screen "参数修改画面" 1280x733, template "模板_2"
   on GenerateScreen: function_b456aad1(1, N); SetTag("变量_100", 17)
   TextField "文本域_7" at 30,0 size 574x42; Text '出现保养提示，请在 查看 / 유지보수 알림이 표시되면, 에서 확인하세요.'
      Visibility <- "VBS_maintenanceWarnStatus_index"
   Button "按钮_4" at 326,0 size 140x42; TextOff '自动画面 / 自動画面: / 자동화면'
      on Press: ActivateScreen("自动画面", 0)
      Visibility <- "VBS_maintenanceWarnStatus_index"
   TextField "文本域_8" at 30,0 size 714x42; Text '保养提示已隐藏，请在 查看 / 유지보수 알림 이미 숨김 , 에서 확인하세요.'
      Visibility <- "VBS_alwaysFalse"
   Button "按钮_3" at 352,0 size 168x42; TextOff '自动画面 / 自動画面: / 자동화면'
      on Press: ActivateScreen("自动画面", 0)
      Visibility <- "VBS_alwaysFalse"
   IOField "IO Field_1" at 195,85 size 121x40; FormatPattern 999
      ProcessValue <- "ST_HMI_Var_HMI_r64NianDu_QianShen_Best"
   TextField "Text Field_13" at 328,155 size 70x32; Text 'mm/s'
   IOField "IO Field_7" at 195,151 size 121x40; FormatPattern 9999
      ProcessValue <- "ST_HMI_Var_HMI_r64Velocity_ChuChe"
   TextField "Text Field_4" at 21,157 size 170x31; Text '出车速度: / 出機速度: / 외진속도:'
   TextField "Text Field_3" at 15,85 size 176x38; Text '牵伸捻度匹配值: ドラフト撚数マッチン グ値: 트위스트 연도 매칭값:'
   TextField "Text Field_9" at 21,216 size 170x38; Text '追捻开始捻度: 追撚開始撚数: 헤드 트위스트 시작 연도:'
   IOField "IO Field_4" at 195,216 size 121x40; FormatPattern 9999
      ProcessValue <- "ST_HMI_Var_HMI_r64NianDu_1"
      ObjectEnable <- "ST_HMI_Var_HMI_boNianDu_3"
   TextField "Text Field_10" at 328,220 size 70x32; Text 'T/M'
   TextField "Text Field_11" at 328,285 size 70x32; Text 'r/min'
   IOField "IO Field_5" at 195,282 size 121x40; FormatPattern 99999
      ProcessValue <- "ST_HMI_Var_HMI_r64NianSu_2"
   TextField "Text Field_24" at 15,282 size 176x38; Text '追捻锭子速度: 追撚スピンドル回転数: 헤드 트위스트 스핀들 속도:'
   TextField "Text Field_29" at 392,25 size 94x30; Text '支数: / 番手: / 번수:'
   IOField "IO Field_18" at 488,20 size 121x40; FormatPattern 99.9
      ProcessValue <- "ST_HMI_Var_HMI_r64ZhiShu_ChengSha"
   TextField "Text Field_2" at 21,25 size 170x31; Text '总捻度: / 総撚数: / 전체 연도:'
   TextField "Text Field_6" at 328,25 size 70x32; Text 'T/M'
   IOField "IO Field_43" at 195,20 size 121x40; FormatPattern 9999
      ProcessValue <- "ST_HMI_Var_HMI_r64NianDu_all"
   TextField "Text Field_7" at 615,23 size 60x32; Text 'Nm'
   Button "按钮_2" at 374,441 size 169x69; TextOn '启用按下 / 使用 / 작동 클릭:'; TextOff '启用 / 使用 / 사용'
      on Press: function_bbf3fe93(1, N)
      on Change: SetBit("ST_Calculation_Var_HMI_bo_Calculation_0_Start"); SetTag("ST_Calculation_Var_g_i16_Calculation_0_3_Select_Status", 1)
      on Release: SetBit("ST_Calculation_Var_HMI_bo_Calculation_0_Start"); SetTag("ST_Calculation_Var_g_i16_Calculation_0_3_Select_Status", 1)
   TextField "Text Field_15" at 615,155 size 60x32; Text 'r/min'
   IOField "IO Field_2" at 488,151 size 121x40; FormatPattern 99999
      ProcessValue <- "ST_HMI_Var_HMI_r64NianSu_Max"
      Appearance <- "ST_HMI_Var_HMI_boAlarm_NianDu_Time"
   IOField "IO Field_13" at 488,85 size 121x40; FormatPattern 99.9
      ProcessValue <- "ST_HMI_Var_HMI_r64Time_JiaNian"
      Appearance <- "ST_HMI_Var_HMI_boAlarm_NianDu_Time"
   TextField "Text Field_48" at 615,89 size 52x32; Text 's'
   Button "按钮_5" at 374,594 size 169x69; TextOn '返回 / リターン / 리턴'; TextOff '返回 / リターン / 리턴'
      on Release: ActivateScreen("设置画面", 0)
   Button "按钮_1" at 1106,176 size 145x54; TextOff '返回 / リターン / 리턴'
      on Click: ActivateScreen("设置画面", 0)
   TextField "Text Field_16" at 690,20 size 142x38; Text '捻缩捻度: ジャッキング．イン 開始撚数: 연축거리:'
   TextField "Text Field_20" at 690,85 size 142x38; Text '捻缩距离: ジャッキング．イン 距離: 연축 트위스트:'
   TextField "Text Field_17" at 970,24 size 63x32; Text 'T/M'
   TextField "Text Field_33" at 970,89 size 63x32; Text 'mm'
   IOField "IO Field_3" at 839,20 size 121x40; FormatPattern 9999
      ProcessValue <- "ST_HMI_Var_HMI_r64NianDu_NianSuo"
   IOField "IO Field_6" at 839,85 size 121x40; FormatPattern 999
      ProcessValue <- "ST_HMI_Var_HMI_r64Position_NianSuo"
      Appearance <- "ST_HMI_Var_HMI_boAlarm_NianSuo_PosNon"
   Button "OBJECT_107" at 400,216 size 232x40; TextOn '追捻启用 / 追撚使用 / 헤드 트위스트 사용'; TextOff '追捻启用 / EXIT / 追撚使用 / 헤드 트위스트 사용'
      on Release: SetBit("ST_HMI_Var_HMI_boNianDu_3")
      Appearance <- "ST_HMI_Var_HMI_boNianDu_3"
   Button "OBJECT_1" at 400,280 size 232x40; TextOn '追捻停用 / 追撚停止 / 헤드 트위스트 사용중지'; TextOff '追捻停用 / EXIT / 追撚停止 / 헤드 트위스트 사용중지'
      on Release: ResetBit("ST_HMI_Var_HMI_boNianDu_3"); SetTag("ST_HMI_Var_HMI_r64NianDu_1", "ST_HMI_Var_HMI_r64NianDu_all")
      Appearance <- "ST_HMI_Var_HMI_boNianDu_3"
   TextField "Text Field_34" at 970,154 size 63x33; Text 's'
   TextField "Text Field_18" at 392,85 size 94x38; Text '加捻时间: / 撚掛時間: / 연사시간:'
   TextField "Text Field_19" at 392,151 size 94x38; Text '锭子速度: スピンドル 回転数: 스핀들속도:'
   Button "按钮_6" at 672,440 size 169x69; TextOn '启用按下 / 使用 / 작동 클릭:'; TextOff '启用 / 使用 / 사용'; TextList "g_i16_Calculation_0_Status"
      Appearance <- "ST_Calculation_Var_g_i16_Calculation_0_Status"
      ProcessValue <- "ST_Calculation_Var_g_i16_Calculation_0_Status"
   TextField "Text Field_14" at 600,533 size 170x31; Text '生效总捻度: / 総撚数: / 전체 연도:'
   TextField "Text Field_23" at 600,600 size 170x31; Text '生效支数: / 総撚数: / 전체 연도:'
   TextField "Text Field_1" at 40,392 size 256x32; Text '更改参数步骤： / パラメーター変更手順: / 매개변수 변경 순서:'
   TextField "Text Field_8" at 38,445 size 277x32; Text '1.更改参数 / １．パラメーター変更 / 1.매개변수 변경'
   TextField "Text Field_12" at 38,510 size 277x32; Text '2.点击“启用” / ２．「使用」をクリック / 2.“사용”을 클릭'
   TextField "Text Field_5" at 38,575 size 277x32; Text '3.点击“返回” / ３．「リターン」をクリック / 3.리턴을 클릭'
   TextField "Text Field_21" at 695,150 size 137x38; Text '捻缩时间: ジャッキング．イン 時間: 연축시간:'
   TextField "Text Field_22" at 695,215 size 137x38; Text '捻缩速度: ジャッキング．イン 速度: 연축속도:'
   TextField "Text Field_31" at 695,285 size 137x32; Text '卷绕长度: / 巻取長: / 와인딩 길이:'
   TextField "Text Field_35" at 970,219 size 63x32; Text 'mm/s'
   TextField "Text Field_36" at 970,285 size 63x32; Text 'mm'
   IOField "IO Field_11" at 839,150 size 121x40; FormatPattern 99.9
      ProcessValue <- "ST_HMI_Var_HMI_r64Time_NianSuo"
   IOField "IO Field_12" at 839,215 size 121x40; FormatPattern 99.9
      ProcessValue <- "ST_HMI_Var_HMI_r64Velocity_NianSuo"
      Appearance <- "ST_HMI_Var_HMI_boAlarm_NianSuo_SuDuOver"
   IOField "IO Field_19" at 839,281 size 121x40; FormatPattern 9999
      ProcessValue <- "ST_HMI_Var_HMI_r64Length_JuanRao"
   IOField "IO Field_8" at 784,600 size 121x40; FormatPattern 99.9
      ProcessValue <- "ST_1TCP_g_myStructSend__lreal_20"
   IOField "IO Field_9" at 784,528 size 121x40; FormatPattern 9999
      ProcessValue <- "ST_1TCP_g_myStructSend__lreal_1"

screen "配方保存画面" 1280x733, template "模板_2"
   on GenerateScreen: function_b456aad1(1, N); SetTag("变量_100", 19)
   TextField "文本域_7" at 30,0 size 574x42; Text '出现保养提示，请在 查看 / 유지보수 알림이 표시되면, 에서 확인하세요.'
      Visibility <- "VBS_maintenanceWarnStatus_index"
   Button "按钮_4" at 326,0 size 140x42; TextOff '自动画面 / 自動画面 / 자동화면'
      on Press: ActivateScreen("自动画面", 0)
      Visibility <- "VBS_maintenanceWarnStatus_index"
   TextField "文本域_8" at 30,0 size 574x42; Text '保养提示已隐藏，请在 查看 / 유지보수 알림 이미 숨김 , 에서 확인하세요.'
      Visibility <- "VBS_alwaysFalse"
   Button "按钮_3" at 352,0 size 168x42; TextOff '自动画面 / 自動画面 / 자동화면'
      on Press: ActivateScreen("自动画面", 0)
      Visibility <- "VBS_alwaysFalse"
   IOField "IO Field_1" at 198,85 size 121x40; FormatPattern 999
      on OnFinishInput: SetBit("ST_Calculation_Var_HMI_bo_Calculation_0_Start"); SetTag("ST_Calculation_Var_g_i16_Calculation_0_3_Select_Status", 1)
      ProcessValue <- "ST_HMI_Var_HMI_r64NianDu_QianShen_Best"
   TextField "Text Field_13" at 331,155 size 70x32; Text 'mm/s'
   IOField "IO Field_7" at 198,151 size 121x40; FormatPattern 9999
      on OnFinishInput: SetBit("ST_Calculation_Var_HMI_bo_Calculation_0_Start"); SetTag("ST_Calculation_Var_g_i16_Calculation_0_3_Select_Status", 1)
      ProcessValue <- "ST_HMI_Var_HMI_r64Velocity_ChuChe"
   TextField "Text Field_4" at 24,157 size 170x31; Text '出车速度: / 出機速度: / 외진속도:'
   TextField "Text Field_3" at 18,85 size 176x38; Text '牵伸捻度匹配值: ドラフト撚数マッチン グ値: 트위스트 연도 매칭값:'
   TextField "Text Field_9" at 24,216 size 170x38; Text '追捻开始捻度: 追撚開始撚数: 헤드 트위스트 시작 연도:'
   IOField "IO Field_4" at 198,216 size 121x40; FormatPattern 9999
      on OnFinishInput: SetBit("ST_Calculation_Var_HMI_bo_Calculation_0_Start"); SetTag("ST_Calculation_Var_g_i16_Calculation_0_3_Select_Status", 1)
      ProcessValue <- "ST_HMI_Var_HMI_r64NianDu_1"
      ObjectEnable <- "ST_HMI_Var_HMI_boNianDu_3"
   TextField "Text Field_10" at 331,220 size 70x32; Text 'T/M'
   TextField "Text Field_11" at 331,285 size 70x32; Text 'r/min'
   IOField "IO Field_5" at 198,282 size 121x40; FormatPattern 99999
      on OnFinishInput: SetBit("ST_Calculation_Var_HMI_bo_Calculation_0_Start"); SetTag("ST_Calculation_Var_g_i16_Calculation_0_3_Select_Status", 1)
      ProcessValue <- "ST_HMI_Var_HMI_r64NianSu_2"
   TextField "Text Field_24" at 18,282 size 176x38; Text '追捻锭子速度: 追撚スピンドル回転数: 헤드 트위스트 스핀들 속도:'
   TextField "Text Field_29" at 366,25 size 101x30; Text '支数: / 番手: / 번수:'
   IOField "IO Field_18" at 469,20 size 121x40; FormatPattern 99.9
      ProcessValue <- "ST_HMI_Var_HMI_r64ZhiShu_ChengSha"
   TextField "Text Field_2" at 24,25 size 170x31; Text '总捻度: / 総撚数: / 전체 연도:'
   TextField "Text Field_6" at 331,25 size 70x32; Text 'T/M'
   IOField "IO Field_43" at 198,20 size 121x40; FormatPattern 9999
      on OnFinishInput: SetBit("ST_Calculation_Var_HMI_bo_Calculation_0_Start"); SetTag("ST_Calculation_Var_g_i16_Calculation_0_3_Select_Status", 1)
      ProcessValue <- "ST_HMI_Var_HMI_r64NianDu_all"
   TextField "Text Field_7" at 596,23 size 60x32; Text 'Nm'
   Button "按钮_5" at 1067,584 size 169x69; TextOff '删除数据记录 / 保存データの削除 / 데이터 기록 삭제'
      on Click: function_be763222("配方视图_1")
   Button "按钮_1" at 680,584 size 169x69; TextOff '当前值显示 / 目前値表示 / 현재값 표시'
      on Click: function_b9843780("配方视图_1")
   Button "按钮_7" at 1107,191 size 145x54; TextOff '返回 / リターン / 리턴'
      on Click: ActivateScreen("设置画面", 0)
   Button "按钮_2" at 861,584 size 193x69; TextOff '数据记录另存为 データを新たに保存する 데이터 기록을 다른 이름으로 저장'
      on Click: function_f5cdec3f("配方视图_1")
   IOField "IO Field_3" at 839,20 size 121x40; FormatPattern 9999
      ProcessValue <- "ST_HMI_Var_HMI_r64NianDu_NianSuo"
   IOField "IO Field_6" at 839,85 size 121x40; FormatPattern 999
      ProcessValue <- "ST_HMI_Var_HMI_r64Position_NianSuo"
   Button "OBJECT_107" at 400,216 size 232x40; TextOn '追捻启用 / 追撚使用 / 헤드 트위스트 사용'; TextOff '追捻启用 / EXIT / 追撚使用 / 헤드 트위스트 사용'
      on Release: SetBit("ST_HMI_Var_HMI_boNianDu_3")
      on Change: SetBit("ST_Calculation_Var_HMI_bo_Calculation_0_Start"); SetTag("ST_Calculation_Var_g_i16_Calculation_0_3_Select_Status", 1)
      Appearance <- "ST_HMI_Var_HMI_boNianDu_3"
   Button "OBJECT_1" at 400,280 size 232x40; TextOn '追捻停用 / 追撚停止 / 헤드 트위스트 사용중지'; TextOff '追捻停用 / EXIT / 追撚停止 / 헤드 트위스트 사용중지'
      on Release: ResetBit("ST_HMI_Var_HMI_boNianDu_3"); SetTag("ST_HMI_Var_HMI_r64NianDu_1", "ST_HMI_Var_HMI_r64NianDu_all")
      on Change: SetBit("ST_Calculation_Var_HMI_bo_Calculation_0_Start"); SetTag("ST_Calculation_Var_g_i16_Calculation_0_3_Select_Status", 1)
      Appearance <- "ST_HMI_Var_HMI_boNianDu_3"
   RecipeView "配方视图_1" at 681,376 size 555x188; DataRecordNrCaption '编号: / Nr.: / No.: / N.º: / N°: / 番号: / 번호: / Nr. / №:'; RecipeNameCaption '配方组名称： / Recipe Name: / レシピグループ名称: / 래서피 이름: / Reseptnavn: / Имя рецепта:'; DataRecordNameCaption '子配方名称： / Datensatzname: / Data Record Name: / Nombre de registro: / Nom d'enregistrement : / Nome del set di dati: / レシピ名称: / 데이터 레코드 이름: / Datapostnavn: / Имя блока данных:'
   TextField "Text Field_1" at 26,389 size 235x32; Text '配方保存步骤： / レシピ保存手順: / 레시피 저장 순서:'
   TextField "Text Field_8" at 23,495 size 609x32; Text '2.点击“当前值显示” / ２．「目前値表示」をクリックする / 2.“현재값 표시”를 클릭'
   TextField "Text Field_12" at 23,435 size 609x32; Text '1.选择“配方组名称” / １．「レシピグループ名称」を選択する / 1.“레시피 그룹 명칭”을 선택'
   TextField "Text Field_14" at 23,556 size 609x32; Text '3.点击“数据记录另存为” / ３．「データを新たに保存する」を選択する / 3.“데이터 기록을 다른 이름으로 저장”을 클릭'
   TextField "Text Field_15" at 23,617 size 609x63; Text '4.输入数据记录名：格式为“序号-捻度-支数-年年月月日日” ４．データ名を入力： 順番ー撚数ー番手ー年 月 日 4.데이터 기록명칭을 입력:양식은“순번-연도-번수-년년월월 일일”.'
   TextField "Text Field_16" at 97,663 size 609x32; Text '例：“01-590-265-20160811” / 例：「01－590－265－20160811」 / 예시：“01-590-265-20160811”'
   TextField "Text Field_5" at 690,20 size 142x38; Text '捻缩捻度: ジャッキング．イン 開始撚数: 연축속도:'
   TextField "Text Field_17" at 970,24 size 63x32; Text 'T/M'
   TextField "Text Field_20" at 690,85 size 142x38; Text '捻缩距离: ジャッキング．イン 距離: 연축거리:'
   TextField "Text Field_33" at 970,89 size 63x32; Text 'mm'

screen "配方选择画面" 1280x733, template "模板_2"
   on GenerateScreen: SetTag("变量_100", 18)
   TextField "文本域_7" at 30,0 size 574x42; Text '出现保养提示，请在 查看 / 유지보수 알림이 표시되면, 에서 확인하세요.'
      Visibility <- "VBS_maintenanceWarnStatus_index"
   Button "按钮_4" at 326,0 size 140x42; TextOff '自动画面 / 自動画面 / 자동화면'
      on Press: ActivateScreen("自动画面", 0)
      Visibility <- "VBS_maintenanceWarnStatus_index"
   TextField "文本域_8" at 30,0 size 574x42; Text '保养提示已隐藏，请在 查看 / 유지보수 알림 이미 숨김 , 에서 확인하세요.'
      Visibility <- "VBS_alwaysFalse"
   Button "按钮_3" at 352,0 size 168x42; TextOff '自动画面 / 自動画面 / 자동화면'
      on Press: ActivateScreen("自动画面", 0)
      Visibility <- "VBS_alwaysFalse"
   IOField "IO Field_1" at 204,85 size 121x40; FormatPattern 999
      on OnFinishInput: SetBit("ST_Calculation_Var_HMI_bo_Calculation_0_Start"); SetTag("ST_Calculation_Var_g_i16_Calculation_0_3_Select_Status", 1)
      ProcessValue <- "ST_HMI_Var_HMI_r64NianDu_QianShen_Best"
   TextField "Text Field_13" at 337,155 size 70x32; Text 'mm/s'
   IOField "IO Field_7" at 204,151 size 121x40; FormatPattern 9999
      on OnFinishInput: SetBit("ST_Calculation_Var_HMI_bo_Calculation_0_Start"); SetTag("ST_Calculation_Var_g_i16_Calculation_0_3_Select_Status", 1)
      ProcessValue <- "ST_HMI_Var_HMI_r64Velocity_ChuChe"
   TextField "Text Field_4" at 24,157 size 176x31; Text '出车速度: / 出機速度: / 외진속도:'
   TextField "Text Field_3" at 24,91 size 176x38; Text '牵伸捻度匹配值: ドラフト撚数マッチン グ値: 트위스트 연도 매칭값:'
   TextField "Text Field_9" at 24,216 size 176x38; Text '追捻开始捻度: 追撚開始撚数: 헤드 트위스트 시작 연도:'
   IOField "IO Field_4" at 204,216 size 121x40; FormatPattern 9999
      on OnFinishInput: SetBit("ST_Calculation_Var_HMI_bo_Calculation_0_Start"); SetTag("ST_Calculation_Var_g_i16_Calculation_0_3_Select_Status", 1)
      ProcessValue <- "ST_HMI_Var_HMI_r64NianDu_1"
   TextField "Text Field_10" at 337,220 size 70x32; Text 'T/M'
   TextField "Text Field_11" at 337,285 size 70x32; Text 'r/min'
   IOField "IO Field_5" at 204,282 size 121x40; FormatPattern 99999
      on OnFinishInput: SetBit("ST_Calculation_Var_HMI_bo_Calculation_0_Start"); SetTag("ST_Calculation_Var_g_i16_Calculation_0_3_Select_Status", 1)
      ProcessValue <- "ST_HMI_Var_HMI_r64NianSu_2"
   TextField "Text Field_24" at 24,282 size 176x38; Text '追捻锭子速度: 追撚スピンドル回転数: 헤드 트위스트 스핀들 속도:'
   TextField "Text Field_29" at 384,25 size 82x30; Text '支数: / 番手: / 번수:'
   IOField "IO Field_18" at 468,20 size 121x40; FormatPattern 99.9
      ProcessValue <- "ST_HMI_Var_HMI_r64ZhiShu_ChengSha"
   TextField "Text Field_2" at 24,25 size 176x31; Text '总捻度: / 総撚数 / 전체 연도:'
   TextField "Text Field_6" at 337,25 size 70x32; Text 'T/M'
   IOField "IO Field_43" at 204,20 size 121x40; FormatPattern 9999
      on OnFinishInput: SetBit("ST_Calculation_Var_HMI_bo_Calculation_0_Start"); SetTag("ST_Calculation_Var_g_i16_Calculation_0_3_Select_Status", 1)
      ProcessValue <- "ST_HMI_Var_HMI_r64NianDu_all"
   TextField "Text Field_7" at 595,23 size 60x32; Text 'Nm'
   Button "按钮_1" at 681,580 size 169x69; TextOff '启用当前配方 / 目前レシピの使用 / 현재 레시피 사용'
      on Click: function_ac24277f("配方视图_1")
      on Release: SetBit("ST_Calculation_Var_HMI_bo_Calculation_0_Start"); SetTag("ST_Calculation_Var_g_i16_Calculation_0_3_Select_Status", 1)
   Button "按钮_7" at 1106,176 size 145x54; TextOff '返回 / リターン / 리턴'
      on Click: ActivateScreen("设置画面", 0)
   RecipeView "配方视图_1" at 681,376 size 555x188; DataRecordNrCaption '编号: / Nr.: / No.: / N.º: / N°: / 番号: / 번호: / Nr. / №:'; RecipeNameCaption '配方组名称： / Recipe Name: / レシピグループ名称: / 래서피 이름: / Reseptnavn: / Имя рецепта:'; DataRecordNameCaption '子配方名称： / Datensatzname: / Data Record Name: / Nombre de registro: / Nom d'enregistrement : / Nome del set di dati: / レシピ名称: / 데이터 레코드 이름: / Datapostnavn: / Имя блока данных:'
   TextField "Text Field_1" at 40,389 size 227x32; Text '配方选择步骤： / レシピ選択手順: / 레시피 선택 순서:'
   TextField "Text Field_8" at 39,495 size 592x32; Text '2.选择“子配方名称” / ２．「レシピ名称」を選択する / 2. “하위 레시비 명칭”을 선택'
   TextField "Text Field_12" at 39,435 size 592x32; Text '1.选择“配方组名称” / １．「レシピグループ名称」を選択する / 1.“레시피 그룹 명칭”을 선택'
   TextField "Text Field_14" at 39,556 size 592x32; Text '3.点击“启用当前配方” / ３．「目前レシピ使用」をクリックする / 3. “현재 레시피 사용”을 클릭한다.'
   IOField "IO Field_9" at 839,20 size 121x40; FormatPattern 9999
      on OnFinishInput: SetBit("ST_Calculation_Var_HMI_bo_Calculation_0_Start"); SetTag("ST_Calculation_Var_g_i16_Calculation_0_3_Select_Status", 1)
      ProcessValue <- "ST_HMI_Var_HMI_r64NianDu_NianSuo"
   IOField "IO Field_10" at 839,85 size 121x40; FormatPattern 999
      on OnFinishInput: SetBit("ST_Calculation_Var_HMI_bo_Calculation_0_Start")
      Appearance <- "ST_HMI_Var_HMI_boAlarm_NianSuo_PosNon"
      ProcessValue <- "ST_HMI_Var_HMI_r64Position_NianSuo"
   TextField "Text Field_5" at 698,24 size 140x38; Text '捻缩捻度: ジャッキング．イン 開始撚数: 연축 트위스트:'
   TextField "Text Field_17" at 970,24 size 63x32; Text 'T/M'
   TextField "Text Field_20" at 700,89 size 130x38; Text '捻缩距离: ジャッキング．イン 距離: 연축거리:'
   TextField "Text Field_33" at 970,89 size 63x32; Text 'mm'

screen "常用调试画面" 1280x733
   on GenerateScreen: SetTag("变量_100", 10)
   Button "HmiScreenItemData_1" at 1105,71 size 145x54; TextOn '向后 / Back / 後向き / 뒤로'; TextOff '向后 / Back / 後向き / 뒤로'
      on Release: ActivateScreen("设置画面", 0)
   IOField "IO Field_38" at 730,162 size 112x42; FormatPattern 999
      ProcessValue <- "ST_HMI_Var_HMI_r64Axis_ZouChe_Position_KongDing_12"
   IOField "IO Field_41" at 730,54 size 112x42; FormatPattern 99
      ProcessValue <- "ST_HMI_Var_HMI_r64_MaoZhou_TouShu"
   IOField "IO Field_10" at 730,108 size 112x42; FormatPattern 999.9
      ProcessValue <- "ST_HMI_Var_HMI_r64Axis_ZouChe_Position_ShengTou_Start_Position"
   IOField "IO Field_28" at 100,322 size 108x40; FormatPattern 99.99
      ProcessValue <- "ST_HMI_Var_HMI_r64_k_ZhangLi_Rate"
   IOField "IO Field_21" at 100,270 size 108x41; FormatPattern 99.99
      ProcessValue <- "ST_HMI_Var_HMI_g1_n_delt_new_0"
   IOField "IO Field_20" at 100,216 size 108x41; FormatPattern 99.99
      ProcessValue <- "ST_HMI_Var_HMI_f1_n_delt_new_0"
   IOField "IO Field_22" at 100,163 size 108x40; FormatPattern 99.99
      ProcessValue <- "ST_HMI_Var_HMI_r64Axis_1_ZhangLi_Position_JuanRao_Set_N"
   IOField "IO Field_23" at 100,109 size 108x40; FormatPattern 99.99
      ProcessValue <- "ST_HMI_Var_HMI_r64Axis_1_ZhangLi_Position_JuanRao_Set_ND"
   IOField "IO Field_24" at 100,55 size 108x40; FormatPattern 99.99
      ProcessValue <- "ST_HMI_Var_HMI_r64Axis_1_ZhangLi_Position_JuanRao_Set_0"
   IOField "IO Field_57" at 100,427 size 109x41; FormatPattern 9.99
      ProcessValue <- "ST_HMI_Var_HMI_k_TuiRao"
   IOField "IO Field_58" at 100,480 size 109x41; FormatPattern 9.99
      ProcessValue <- "ST_HMI_Var_HMI_scalevalue_Cam_3"
   IOField "IO Field_1" at 100,594 size 108x40; FormatPattern 99999
      ProcessValue <- "ST_Main_Var_g_r64Axis_DingZi_PositiveAccel_CunRao"
   IOField "IO Field_25" at 100,648 size 108x40; FormatPattern 99.99
      ProcessValue <- "ST_Main_Var_g_r64Axis_DingZi_Velocity_CunRao_ratio"
   Button "HmiScreenItemData_2" at 1104,352 size 145x54; TextOn '向后 / 後向き / 뒤로'; TextOff '张力测定 / 張力測定 / 장력 측정'; Authorization "Operate_4"
      on Release: ActivateScreen("张力测定", 0)
   Button "HmiScreenItemData_3" at 1104,424 size 145x54; TextOn '向后 / 後向き / 뒤로'; TextOff '原点设定 / 原点設定 / 원점 설정'; Authorization "Operate_4"
      on Release: ActivateScreen("原点设定", 0)
   Button "HmiScreenItemData_4" at 1104,496 size 145x54; TextOn '向后 / 後向き / 뒤로'; TextOff '纱管参数设定 糸管パラメーター 設定 보빈 매개변수 설정'; Authorization "Operate_4"
      on Release: ActivateScreen("纱管参数设定", 0)
   Button "Template_Button_1" at 791,673 size 85x59; TextOff 'Text'; PictureOff "China_1"
      on Click: function_fb9197e8(-1)
   Button "HmiScreenItemData_15" at 928,679 size 158x53; TextOn '6卷绕相关1 / 6巻取関係1'; TextOff '校准触摸屏 / タッチパネルの校正 / 터치 스크린 교정'
      on Release: function_bc3e350c()
   IOField "IO Field_2" at 729,214 size 112x42; FormatPattern 99.9
      ProcessValue <- "ST_HMI_Var_HMI_r64Axis_ZouChe_Position_ZiDongTingZhi"
   IOField "IO Field_3" at 729,270 size 112x42; FormatPattern 999
      ProcessValue <- "ST_HMI_Var_HMI_r64Axis_ZouChe_Position_ChuChe_Middle"
   Button "HmiScreenItemData_6" at 1104,570 size 145x54; TextOn '向后 / 後向き / 뒤로'; TextOff '纱穗参数设定 糸管パラメーター 設定 코프 매개변수'; Authorization "Operate_4"
      on Release: ActivateScreen("纱穗参数设定", 0)
   IOField "IO Field_8" at 728,392 size 112x42; FormatPattern 99999
      Visibility <- "ST_Calculation_Var_Date_Temp"
      ProcessValue <- "ST_Calculation_Var_g_r64Axis_DingZi_PositiveAccel_Buffer_JiaNian{1}"
      Appearance <- "ST_HMI_Var_HMI_boAlarm_NianDu_Time"
   IOField "IO Field_7" at 728,392 size 112x42; FormatPattern 99999
      Visibility <- "ST_Calculation_Var_Date_Temp"
      ProcessValue <- "ST_Calculation_Var_g_r64Axis_DingZi_PositiveAccel_Buffer_JiaNian{0}"
      Appearance <- "ST_HMI_Var_HMI_boAlarm_NianDu_Time"
   Button "Template_Button_11" at 1196,673 size 78x59; TextOn 'NavigateHome'; TextOff 'NavigateHome'; PictureOn "NavigateHome_TP1200_Comfort"; PictureOff "NavigateHome_TP1200_Comfort"
      on Release: ActivateScreen("自动画面", 0); function_f23ef4c9()
   TextField "Text Field_44" at 219,427 size 290x41; Text '退绕曲线拐点比例 / パッキングオフ湾曲点比例 / 언와인딩 곡선 변곡점 비율'
   TextField "Text Field_46" at 219,480 size 254x41; Text '退绕圈数比例 / パッキングオフ巻取比例 / 언와인딩 랩수 비율'
   TextField "Text Field_37" at 222,218 size 430x41; Text '卷绕速度中点调整值—初始值 / 中間点の取り巻き速度調整値ー初期値 / 와인딩 속도 중심점조정값-초기값'
   TextField "Text Field_38" at 222,272 size 430x41; Text '卷绕速度末点调整值—初始值 / 終了時点の取り巻き速度調整値ー初期値 / 와인딩 속도 종료점조정값-초기값'
   TextField "Text Field_39" at 222,165 size 430x41; Text '卷绕张力弓目标值—满纱时 / カウンターフォーラーの目標値ー満巻時 / 와인딩 장력 호랑 목표값-만사일시'
   TextField "Text Field_40" at 224,112 size 430x41; Text '卷绕张力弓目标值—最大直径时 / カウンターフォーラーの目標値ー最大直径時 / 와이딩 장력 호랑목표값-최대직경일시'
   TextField "Text Field_41" at 222,57 size 430x41; Text '卷绕张力弓目标值—生头时 / カウンターフォーラーの目標値ー巻始め / 와인딩 장력호랑 목표값-실시작점'
   TextField "Text Field_45" at 222,324 size 430x41; Text '卷绕张力弓反馈增益 / カウンターフォーラーのフィードバック増幅 / 와인딩 장력호랑 피드백 게인'
   TextField "Text Field_1" at 222,592 size 430x41; Text '存绕锭子加速度 / 逆巻取スピンドル加速度 / 와인딩 스핀들 가속'
   TextField "Text Field_42" at 222,646 size 430x41; Text '存绕锭子速度比例 / 逆巻取スピンドル回転速度比例 / 와인딩 스핀들 속도 비율'
   TextField "Text Field_58" at 857,164 size 230x41; Text '生头中间停止位置 / 自動停止位置 / 스레딩중 정지위치'
   TextField "Text Field_8" at 857,56 size 230x41; Text '毛轴头数 / 篠棒本数 / 시누 세부샤프트개수'
   TextField "Text Field_2" at 857,110 size 230x41; Text '生头起点位置 / 口付け開始点位置 / 스레딩시작점 위치'
   TextField "Text Field_14" at 100,6 size 233x42; Text '卷绕相关 / 巻取関係 / 와인딩 관련'
   TextField "Text Field_3" at 100,377 size 233x42; Text '退绕相关 / パッキングオフ関連 / 언와인딩 관련'
   TextField "Text Field_4" at 100,542 size 233x42; Text '存绕相关 / 逆巻取関連 / 와인딩관련'
   TextField "Text Field_5" at 778,6 size 233x42; Text '其他 / その他 / 기타'
   Button "按钮_1" at 1104,280 size 145x54; TextOff '牵伸调整 / 연신조절'; Authorization "Operate_4"
      on Press: ActivateScreen("牵伸调整画面", 0)
   TextField "Text Field_6" at 856,216 size 230x41; Text '自动停止位置 / 自動停止位置 / 자동정지위치'
   TextField "Text Field_7" at 856,272 size 230x41; Text '出车停止位置 / 自動停止位置 / 외진정지위치'
   IOField "IO Field_4" at 728,452 size 112x42; FormatPattern 9.99
      on OnFinishInput: SetBit("ST_Calculation_Var_HMI_bo_Calculation_0_Start"); SetTag("ST_Calculation_Var_g_i16_Calculation_0_3_Select_Status", 1)
      ProcessValue <- "ST_TO_DZ_FU_Var_HMI_r64Ratio_PositiveAccelStartJerk_JiaNian"
   IOField "IO Field_6" at 728,508 size 112x42; FormatPattern 9.99
      on OnFinishInput: SetBit("ST_Calculation_Var_HMI_bo_Calculation_0_Start"); SetTag("ST_Calculation_Var_g_i16_Calculation_0_3_Select_Status", 1)
      ProcessValue <- "ST_TO_DZ_FU_Var_HMI_r64Ratio_PositiveAccelEndJerk_JiaNian"
   IOField "IO Field_9" at 728,560 size 112x42; FormatPattern 99.99
      ProcessValue <- "ST_HMI_Var_HMI_r64_DingZi_Zouche_ratio_KongDing_65_1"
   TextField "Text Field_12" at 856,392 size 230x41; Text '锭子加速度'
   TextField "Text Field_9" at 856,448 size 230x41; Text '锭子+Jerk比例'
   TextField "Text Field_11" at 856,504 size 230x41; Text '锭子-Jerk比例'
   TextField "Text Field_13" at 856,560 size 230x41; Text '光锭卷绕传动比1'
   IOField "IO Field_5" at 728,320 size 112x42; FormatPattern 9.99
      on OnFinishInput: SetBit("ST_Calculation_Var_HMI_bo_Calculation_0_Start"); SetTag("ST_Calculation_Var_g_i16_Calculation_0_3_Select_Status", 1)
      ProcessValue <- "ST_HMI_Var_HMI_r64Ratio_PositiveAccel_Jerk_JiaNian"
   TextField "Text Field_10" at 856,320 size 230x41; Text '锭子加速度比例 / 自動停止位置 / 외진정지위치'
   Button "按钮_3" at 1104,208 size 145x54; TextOff '卷绕调整 / 牵伸调整 / 연신조절'; Authorization "Operate_4"
      on Press: ActivateScreen("卷绕经验参数", 0)
   Button "HmiScreenItemData_12" at 1105,138 size 146x52; TextOn '11生头相关'; TextOff '生头相关'; Authorization "Operate_4"
      on Release: ActivateScreen("生头相关", 0)
   Button "Template_Button_2" at 667,673 size 78x59; TextOff 'Text'; PictureOff "1"
      on Click: StopRuntime(0)

screen "张力测定" 1280x733, template "模板_2"
   on GenerateScreen: SetTag("变量_100", 12)
   Button "OBJECT_109" at 120,48 size 182x70; TextOn '张力测定 / 張力測定 / 장력 측정'; TextOff '张力测定 / EXIT / 張力測定 / 장력 측정'
      on Press: SetTag("ST_Main_Var_g_i16_Mode_Selected", 256)
      Appearance <- "ST_Main_Var_g_bo_Mode_Enabled_Manual"
   Button "OBJECT_110" at 120,234 size 182x70; TextOff '张力测定启动 / EXIT / 張力測定起動 / 장력 측정 시작'
      on Release: ResetBit("ST_HMI_Var_HMI_bo_ZhangLi_CeDing_Start")
      on Press: SetBit("ST_HMI_Var_HMI_bo_ZhangLi_CeDing_Start")
      Appearance <- "ST_Main_Var_g_bo_Mode_Enabled_Manual"
   IOField "I/O 域_1" at 502,42 size 86x40; FormatPattern 99.99
      ProcessValue <- "ST_Var_ZLCD_HMI_r64Axis_1_ZhangLi_Torque_CeDing_N{0}"
   IOField "I/O 域_2" at 502,86 size 86x40; FormatPattern 99.99
      ProcessValue <- "ST_Var_ZLCD_HMI_r64Axis_1_ZhangLi_Torque_CeDing_N{1}"
   IOField "I/O 域_3" at 502,130 size 86x40; FormatPattern 99.99
      ProcessValue <- "ST_Var_ZLCD_HMI_r64Axis_1_ZhangLi_Torque_CeDing_N{2}"
   IOField "I/O 域_4" at 502,174 size 86x40; FormatPattern 99.99
      ProcessValue <- "ST_Var_ZLCD_HMI_r64Axis_1_ZhangLi_Torque_CeDing_N{3}"
   IOField "I/O 域_5" at 502,218 size 86x40; FormatPattern 99.99
      ProcessValue <- "ST_Var_ZLCD_HMI_r64Axis_1_ZhangLi_Torque_CeDing_N{4}"
   IOField "I/O 域_6" at 502,261 size 86x40; FormatPattern 99.99
      ProcessValue <- "ST_Var_ZLCD_HMI_r64Axis_1_ZhangLi_Torque_CeDing_N{6}"
   Button "按钮_1" at 726,234 size 182x70; TextOn '调整 / 調整 / 조정'; TextOff '调整 / 調整 / 조정'
      on Release: ResetBit("ST_Var_ZLCD_HMI_bo_ZhangLi_CeDing_Adjustment")
      on Press: SetBit("ST_Var_ZLCD_HMI_bo_ZhangLi_CeDing_Adjustment")
   TextField "文本域_6" at 60,336 size 996x358; Text '张力弓整定步骤 1. 按一下“手动”按钮，按“成形弓降”按钮，将成形钢丝降到锭尖附近，按一下“去使能”按钮 2. 拉住张力弓，同时按住“停止”和“张力弓降”两个按钮，张力电机抱闸会松开电机抱闸，让张 力钢丝掉到走车撞块上 3. 按一下“手动按钮” 4. 点击“张力测定”，点击“张力测定启动” 5. 张力钢丝自动从最低点开始缓慢上升，同时自动记录数据 6. 待上升到48.5左右时张力弓停下 7. 观察以上6个数据，按下右侧的“调整”按钮，可看到前三个数据被第四个覆盖 8. 按下手动——>张力弓降，将张力钢丝降到正常位置 9. 结束 カウンターフォーラー調整手順 １．”手動”を一度押し、”ワイディングフォーラー下降”ボタンを押して”ワイディングフォーラー”ワイヤをスピンド ルの先端までさげ、”長期停止”ボタンを一度押す。 ２．”カウンターフォーラー”を引きながら、同時に”停止”と”カウンターフォーラー下降”ボタンを一度押す。カウ ンターモーターの制動を緩み、”ワイディングフォーラー”ワイヤをキャレージのブロックに落とせる。 ３．一度”手動”ボタンを押す ４．”張力測定”をクリックし、また”張力測定起動”をクリックする。 ５．カウンターワイヤを自動で下死点から徐々に上昇させながら、同時に自動でデータを記録する。 ６．48.5前後に上昇となった時点で、カウンターフォーラーを停止させる。 ７．以上の六つのデータを観察しながら、右側の”調整”ボタンを一度押すと、前の三つのテータが四つ目のデ ータに切り替わったことが分かる。 8．順序に”手動”と”カウンターフォーラー下降”ボタンを押せ、カウンターワイヤをさげる。 9．终。 장력 호랑셋업 순서 1. “수동”버튼을 누르고 “성형호랑하강” 버튼을 눌러 성형호랑 을스핀들 팁 근처까지 내려오게 하고 ‘비활성화’버튼을 누른다. 2. 장력호랑을당기고“정지”와 “장력호랑하강”두 버튼을 동시에 누른다.장력 호랑모터 브레이크가 풀리 면서 장력 와이어가 캐리지링크 스토퍼에 떨어진다. 3. “수동버튼”을 누른다. 4. “장력측정”을클릭하고“장력측정 시작”을 클릭한다. 5. 장력 와이어는 자동으로 최저포인트로부터 시작하여 천천히 상승하면서 자동으로 데이터를 기록한다. 6. 48. 5좌우까지 상승하면 장력 호랑을 정지한다. 7. 이상 6개데이터를 관찰하고 우측의 “조정”버튼을 누르면 처음3개 데이터가 네번째에 의해커버되어 있 는것을 볼수 있다. 8. 수동——>장력 호랑하강을 눌러 장력 와이어를 정상위치까지 내린다. 9. 종료'
   TextField "文本域_1" at 30,541 size 17x21; Text 'Text'
   Button "HmiScreenItemData_2" at 1106,174 size 145x54; TextOn '向后 / 後向き / 뒤로'; TextOff '向后 / 後向き / 뒤로'
      on Release: ActivateScreen("设置画面", 0)
   Button "HmiScreenItemData_3" at 1106,362 size 145x54; TextOn '向后 / 後向き / 뒤로'; TextOff '张力测定 / 張力測定 / 장력 측정'
      on Release: ActivateScreen("张力测定", 0)
   Button "HmiScreenItemData_4" at 1106,452 size 145x54; TextOn '向后 / 後向き / 뒤로'; TextOff '原点设定 / 原点設定 / 원점 설정'
      on Release: ActivateScreen("原点设定", 0)
   Button "HmiScreenItemData_5" at 1106,542 size 145x54; TextOn '向后 / 後向き / 뒤로'; TextOff '纱管参数设定 糸管パラメーター 設定 보빈 매개변수 설정'
      on Release: ActivateScreen("纱管参数设定", 0)
   Button "HmiScreenItemData_6" at 1106,272 size 145x54; TextOn '向后 / 後向き / 뒤로'; TextOff '常用调试画面 / 常用調整画面 / 상용 조정화면'
      on Release: ActivateScreen("常用调试画面", 0)

screen "原点设定" 1280x733, template "模板_2"
   on GenerateScreen: SetTag("变量_100", 13)
   IOField "I/O 域_1" at 885,196 size 88x48; FormatPattern 99
      ProcessValue <- "ST_HMI_Var_HMI_r64StartPosition_Axis_ZouChe_0"
   TextField "文本域_1" at 78,194 size 260x48; Text '走车编码器当前位置 キャレージのエンコー ダーの目前位置 캐리지 인코더 현재 위치'
   IOField "I/O 域_2" at 351,194 size 88x48; FormatPattern 99999.99
      ProcessValue <- "Axis_ZouChe_positioningState_actualPosition"
   Button "按钮_4" at 789,195 size 76x47; TextOff '出车 / 出機 / 외진'
      on Release: ResetBit("ST_HMI_Var_HMI_bo_ChuChe")
      on Press: SetBit("ST_HMI_Var_HMI_bo_ChuChe")
   Button "按钮_5" at 458,194 size 76x47; TextOff '进车 / 入機 / 내진'
      on Release: ResetBit("ST_HMI_Var_HMI_bo_JinChe")
      on Press: SetBit("ST_HMI_Var_HMI_bo_JinChe")
   IOField "I/O 域_3" at 885,304 size 88x48; FormatPattern 99.999
      ProcessValue <- "ST_HMI_Var_HMI_r64StartPosition_Axis_1_ZhangLi_0"
   IOField "I/O 域_4" at 885,413 size 88x48
      ProcessValue <- "ST_HMI_Var_HMI_r64StartPosition_Axis_ChengXing_0"
   TextField "文本域_2" at 78,302 size 260x48; Text '张力编码器当前位置 カウンターのエンコー ダーの目前位置 장력 인코더 현재 위치'
   IOField "I/O 域_5" at 351,302 size 88x48; FormatPattern 999.99
      ProcessValue <- "Axis_1_ZhangLi_positioningState_actualPosition"
   Button "按钮_1" at 789,303 size 76x47; TextOff '升 / 上昇 / 상승'
      on Release: ResetBit("ST_HMI_Var_HMI_bo_ZhangLi_Up")
      on Press: SetBit("ST_HMI_Var_HMI_bo_ZhangLi_Up")
   Button "按钮_2" at 458,302 size 76x47; TextOff '降 / 下降 / 하강'
      on Release: ResetBit("ST_HMI_Var_HMI_bo_ZhangLi_Down")
      on Press: SetBit("ST_HMI_Var_HMI_bo_JinChe")
   TextField "文本域_3" at 78,412 size 260x48; Text '成形编码器当前位置 ワインディングのエンコ ーダーの目前位置 성형 인코더 현재 위치'
   IOField "I/O 域_6" at 351,412 size 88x48; FormatPattern 9999.99
      ProcessValue <- "Axis_ChengXing_positioningState_actualPosition"
   Button "按钮_3" at 458,413 size 76x47; TextOff '升 / 上昇 / 상승'
      on Release: ResetBit("ST_HMI_Var_HMI_bo_ChengXing_Up")
      on Press: SetBit("ST_HMI_Var_HMI_bo_ChuChe")
   Button "按钮_6" at 789,414 size 76x47; TextOff '降 / 下降 / 하강'
      on Release: ResetBit("ST_HMI_Var_HMI_bo_ChengXing_Down")
      on Press: SetBit("ST_HMI_Var_HMI_bo_ChengXing_Down")
   Bar "棒图_1" at 554,195 size 216x49; MinimumValue 40; MaximumValue 90
      ProcessValue <- "Axis_ZouChe_positioningState_actualPosition"
   Bar "棒图_2" at 554,301 size 216x49; MinimumValue 50; MaximumValue 70
      ProcessValue <- "Axis_1_ZhangLi_positioningState_actualPosition"
   Bar "棒图_3" at 554,410 size 216x49; MinimumValue 320; MaximumValue 335
      ProcessValue <- "Axis_ChengXing_positioningState_actualPosition"
   Button "按钮_7" at 56,618 size 280x50; TextOn '微调模式 / 微調整'; TextOff '按下进入微调模式 / 微調整モードに切り替える / 미세조정 모드진입 을 누른다.'
      on Release: ResetBit("ST_HMI_Var_HMI_boMinorAdjustment_select")
      on Press: SetBit("ST_HMI_Var_HMI_boMinorAdjustment_select")
   Button "HmiScreenItemData_2" at 846,683 size 159x48; TextOn '报警画面 / 警報画面 / 경보알람화면'; TextOff '报警画面 / 警報画面 / 경보알람화면'
      on Release: ActivateScreen("报警画面", 0)
   Button "OBJECT_106" at 1039,2 size 238x42; TextOff '手动 / EXIT / 手動 / 수동'; TextList "mode_enabled_1"
      ProcessValue <- "ST_Main_Var_g_i16_Mode_Enabled"
      Appearance <- "ST_Main_Var_g_i16_Mode_Enabled"
   TextField "文本域_6" at 168,88 size 807x58; Text '注意： 不要随意修改此页的数据，不当的数据可能导致行程超限撞车的危险！ 注意：勝手に本ページのデータを変えてはいけない。不当なデータはキャレージのストロー クのオーバーを招き衝突の危険がある。 주의:임의로 이 페이지의 데이터를 수정하지 마십시오.부적절한 데이터는 스트로크 오버런충돌 위험을 초래할수 있습니다!'
   GraphicView "图形视图_2" at 57,70 size 102x99; Picture "图形_2"
   Button "HmiScreenItemData_3" at 1106,174 size 145x54; TextOn '向后 / 後向き / 뒤로'; TextOff '向后 / 後向き / 뒤로'
      on Release: ActivateScreen("设置画面", 0)
   Button "HmiScreenItemData_4" at 1106,362 size 145x54; TextOn '向后 / 後向き / 뒤로'; TextOff '张力测定 / 張力測定 / 장력 측정'
      on Release: ActivateScreen("张力测定", 0)
   Button "HmiScreenItemData_5" at 1106,452 size 145x54; TextOn '向后 / 後向き / 뒤로'; TextOff '原点设定 / 原点設定 / 원점 설정'
      on Release: ActivateScreen("原点设定", 0)
   Button "HmiScreenItemData_6" at 1105,542 size 147x54; TextOn '向后 / 後向き / 뒤로'; TextOff '纱管参数设定 糸管パラメーター 設定 보빈 매개변수 설정'
      on Release: ActivateScreen("纱管参数设定", 0)
   Button "HmiScreenItemData_7" at 1106,272 size 145x54; TextOn '向后 / 後向き / 뒤로'; TextOff '常用调试画面 / 常用調整画面 / 상용 조정화면'
      on Release: ActivateScreen("常用调试画面", 0)

screen "纱管参数设定" 1280x733, template "模板_2"
   on GenerateScreen: SetTag("变量_100", 14)
   IOField "IO Field_41" at 69,59 size 112x42; FormatPattern 99.99
      ProcessValue <- "ST_HMI_Var_HMI_r64_h0_s"
   IOField "IO Field_46" at 69,169 size 112x42; FormatPattern 99.99
      ProcessValue <- "ST_HMI_Var_HMI_r64Diameter_ShaGuan_Middle"
   IOField "IO Field_1" at 69,113 size 112x42; FormatPattern 99.99
      ProcessValue <- "ST_HMI_Var_HMI_r64Diameter_ShaGuan_Bottom"
   IOField "IO Field_2" at 69,279 size 112x42
      ProcessValue <- "ST_HMI_Var_HMI_r64Height_ShaGuan_Middle"
   IOField "IO Field_3" at 69,335 size 112x42
      ProcessValue <- "ST_HMI_Var_HMI_r64Height_ShaGuan_Top"
   IOField "IO Field_6" at 69,223 size 112x42; FormatPattern 99.99
      ProcessValue <- "ST_HMI_Var_HMI_r64Diameter_ShaGuan_Top"
   IOField "IO Field_4" at 69,392 size 112x42; FormatPattern 99.9
      ProcessValue <- "ST_HMI_Var_HMI_r64_DingZi_Zouche_ratio_KongDing_9_Shaguan1"
   IOField "IO Field_5" at 589,59 size 112x42; FormatPattern 99.99
      ProcessValue <- "ST_HMI_Var_HMI_r64_h0_s_2"
   IOField "IO Field_7" at 589,169 size 112x42; FormatPattern 99.99
      ProcessValue <- "ST_HMI_Var_HMI_r64Diameter_ShaGuan_Middle_2"
   IOField "IO Field_8" at 589,113 size 112x42; FormatPattern 99.99
      ProcessValue <- "ST_HMI_Var_HMI_r64Diameter_ShaGuan_Bottom_2"
   IOField "IO Field_9" at 589,279 size 112x42
      ProcessValue <- "ST_HMI_Var_HMI_r64Height_ShaGuan_Middle_2"
   IOField "IO Field_10" at 589,335 size 112x42
      ProcessValue <- "ST_HMI_Var_HMI_r64Height_ShaGuan_Top_2"
   IOField "IO Field_11" at 589,223 size 112x42; FormatPattern 99.99
      ProcessValue <- "ST_HMI_Var_HMI_r64Diameter_ShaGuan_Top_2"
   IOField "IO Field_12" at 589,392 size 112x42; FormatPattern 99.9
      ProcessValue <- "ST_HMI_Var_HMI_r64_DingZi_Zouche_ratio_KongDing_9_Shaguan2"
   TextField "Text Field_8" at 207,59 size 332x42; Text '纱管安装高度 / 糸管装着高度 / 보빈 설치 높이'
   TextField "Text Field_9" at 207,113 size 332x42; Text '纱管底部直径 / 糸管底部直径 / 보빈 하단부분 직경'
   TextField "Text Field_10" at 207,169 size 332x42; Text '纱管中间直径 / 糸管中間部直径 / 보빈 중간부분 직경'
   TextField "Text Field_11" at 207,223 size 332x42; Text '纱管顶部有效直径 / 糸管上部有効直径 / 보빈 상단 유효 직경'
   TextField "Text Field_12" at 207,279 size 332x42; Text '纱管从底部到中间的高度 / 糸管底部から中間部までの高度 / 보빈 하단에서 중간까지의 높이'
   TextField "Text Field_13" at 207,335 size 345x42; Text '纱管从中间到顶部的高度 / 糸管中間部から上部までの高度 / 보빈 중간부분에서 상단까지의 높이'
   TextField "Text Field_1" at 207,392 size 332x42; Text '空锭-锭子走车传动比 / 空鍾－スピンドル キャレージ伝動比 / 아이들 스핀들-스핀들 캐리지 기어비'
   TextField "Text Field_3" at 727,59 size 332x42; Text '纱管安装高度 / 糸管装着高度 / 보빈 설치 높이'
   TextField "Text Field_4" at 727,113 size 332x42; Text '纱管底部直径 / 糸管底部直径 / 보빈 하단부분 직경'
   TextField "Text Field_5" at 727,169 size 332x42; Text '纱管中间直径 / 糸管中間部直径 / 보빈 중간부분 직경'
   TextField "Text Field_6" at 727,223 size 332x42; Text '纱管顶部有效直径 / 糸管上部有効直径 / 보빈 상단 유효 직경'
   TextField "Text Field_7" at 727,279 size 332x42; Text '纱管从底部到中间的高度 / 糸管底部から中間部までの高度 / 보빈 하단에서 중간까지의 높이'
   TextField "Text Field_14" at 727,335 size 345x42; Text '纱管从中间到顶部的高度 / 糸管中間部から上部までの高度 / 보빈 중간부분에서 상단까지의 높이'
   TextField "Text Field_16" at 727,392 size 332x42; Text '空锭-锭子走车传动比 / 空鍾－スピンドル キャレージ伝動比 / 아이들 스핀들-스핀들 캐리지 기어비'
   Button "OBJECT_3" at 69,4 size 160x48; TextOff '标准纱管1： / EXIT / 標準糸管１: / 표준보빈1:'
      on Press: SetTag("ST_HMI_Var_HMI_i16_Status_ShaGuan_Select", 1)
      Appearance <- "ST_HMI_Var_HMI_i16_Status_ShaGuan_Select"
   Button "OBJECT_4" at 589,4 size 160x48; TextOff '标准纱管2： / EXIT / 標準糸管２: / 표준보빈2:'
      on Press: SetTag("ST_HMI_Var_HMI_i16_Status_ShaGuan_Select", 2)
      Appearance <- "ST_HMI_Var_HMI_i16_Status_ShaGuan_Select"
   Button "HmiScreenItemData_2" at 1106,174 size 145x54; TextOn '向后 / 後向き / 뒤로'; TextOff '向后 / 後向き / 뒤로'
      on Release: ActivateScreen("设置画面", 0)
   Button "HmiScreenItemData_3" at 1106,362 size 145x54; TextOn '向后 / 後向き / 뒤로'; TextOff '张力测定 / 張力測定 / 장력 측정'
      on Release: ActivateScreen("张力测定", 0)
   Button "HmiScreenItemData_4" at 1106,452 size 145x54; TextOn '向后 / 後向き / 뒤로'; TextOff '原点设定 / 原点設定 / 원점 설정'
      on Release: ActivateScreen("原点设定", 0)
   Button "HmiScreenItemData_5" at 1106,542 size 145x54; TextOn '向后 / 後向き / 뒤로'; TextOff '纱管参数设定 糸管パラメーター 設定 보빈 매개변수 설정'
      on Release: ActivateScreen("纱管参数设定", 0)
   Button "HmiScreenItemData_6" at 1106,272 size 145x54; TextOn '向后 / 後向き / 뒤로'; TextOff '常用调试画面 / 常用調整画面 / 상용 조정화면'
      on Release: ActivateScreen("常用调试画面", 0)

screen "牵伸调整画面" 1280x733, template "Template"
   on GenerateScreen: SetTag("变量_100", 11)
   IOField "I/O 域_2" at 404,332 size 106x48; FormatPattern 9.999
      ProcessValue <- "ST_HMI_Var_HMI_r64_QianShen_Add1"
   TextField "Text Field_25" at 22,332 size 380x48; Text '牵伸第一次增加量q1： / 연신(드라프트) 제1차 증가량 q1:'
   IOField "I/O 域_1" at 404,414 size 106x48; FormatPattern 9.999
      ProcessValue <- "ST_HMI_Var_HMI_r64_QianShen_Add2"
   TextField "Text Field_1" at 22,414 size 380x48; Text '牵伸第二次增加量q2： / 연신(드라프트) 제2차 증가량 q2:'
   IOField "I/O 域_3" at 404,496 size 106x48; FormatPattern 9999
      ProcessValue <- "ST_HMI_Var_HMI_r64_ShaXian_L1"
   TextField "Text Field_2" at 22,496 size 380x48; Text '牵伸第一次增加时纱线米数L1： 연신(드라프트) 제1차 증가시 원사 메터수 L1:'
   IOField "I/O 域_4" at 404,578 size 106x48; FormatPattern 9999
      ProcessValue <- "ST_HMI_Var_HMI_r64_ShaXian_L2"
   TextField "Text Field_3" at 22,578 size 380x48; Text '牵伸第二次增加时纱线米数L2： 연신(드라프트) 제2차 증가시 원사 메터수 L2:'
   TextField "Text Field_5" at 350,47 size 340x48; Text '牵伸第一次增加量q1： / 연신(드라프트) 제1차 증가량 q1:'
   TextField "Text Field_6" at 700,16 size 340x48; Text '牵伸第二次增加量q2： / 연신(드라프트) 제2차 증가량 q2:'
   TextField "Text Field_7" at 64,0 size 176x48; Text '总牵伸 / 전체 드라프트'
   TextField "Text Field_8" at 1136,207 size 142x48; Text '纱线米数 / 원사 미터수'
   TextField "Text Field_9" at 250,259 size 350x48; Text '牵伸第一次增加时纱线米数L1 연신(드라프트) 제1차 증가시 원사 메터수 L1:'
   TextField "Text Field_10" at 600,259 size 350x48; Text '牵伸第二次增加时纱线米数L2 연신(드라프트) 제2차 증가시 원사 메터수 L2:'
   TextField "Text Field_11" at 1008,259 size 196x48; Text '总纱线米数L3 / 총 원사 미터수 L3'
   IOField "I/O 域_6" at 1125,496 size 106x48; FormatPattern 9.999
      ProcessValue <- "ST_HMI_Var_HMI_r64QianShen_All_real"
   TextField "Text Field_12" at 760,496 size 360x48; Text '实时总牵伸： / 실시간 전체 연신(드라프트):'
   IOField "I/O 域_7" at 1125,332 size 106x48; FormatPattern 9.999
      ProcessValue <- "ST_HMI_Var_HMI_r64QianShen_All"
   TextField "Text Field_13" at 760,332 size 360x48; Text '设置的总牵伸： / 설정한 전체 연신(드라프트):'
   IOField "I/O 域_8" at 1125,414 size 106x48; FormatPattern 9.999
      ProcessValue <- "ST_HMI_Var_HMI_r64QianShen_All_object"
   TextField "Text Field_14" at 760,414 size 360x48; Text '调整后的目标总牵伸： / 조절후의 목표 전체 연신(드라프트):'
   IOField "I/O 域_9" at 610,496 size 106x48; FormatPattern 99
      ProcessValue <- "ST_HMI_Var_HMI_r64_Ratio1"
   IOField "I/O 域_10" at 610,578 size 106x48; FormatPattern 99
      ProcessValue <- "ST_HMI_Var_HMI_r64_Ratio2"
   TextField "Text Field_15" at 491,496 size 119x48; Text '百分比1： / 백분율1:'
   TextField "Text Field_16" at 491,578 size 119x48; Text '百分比2： / 백분율2:'
   TextField "Text Field_4" at 722,496 size 29x48; Text '%'
   TextField "Text Field_17" at 722,578 size 29x48; Text '%'
   Button "HmiScreenItemData_1" at 1072,666 size 159x47; TextOn '向后 / 後向き / 뒤로'; TextOff '向后 / 後向き / 뒤로'
      on Release: ActivateScreen("常用调试画面", 0)

screen "手动画面" 1280x733, template "模板_1"
   on GenerateScreen: SetTag("变量_100", 2)
   Button "HmiScreenItemData_1" at 1119,179 size 159x47; TextOn '向后 / 後向き / 뒤로'; TextOff '向后 / 後向き / 뒤로'
      on Release: ActivateScreen("自动画面", 0)
   Button "HmiScreenItemData_2" at 1119,285 size 159x47; TextOn '手动设置 / 手動設置 / 수동설정'; TextOff '手动设置 / 手動設置 / 수동설정'
      on Release: ActivateScreen("手动设置", 0)
   Button "OBJECT_107" at 873,289 size 177x68; TextOff '去使能 / EXIT / 長期停止 / 비활성화'
      on Release: ResetBit("ST_HMI_Var_HMI_bo_Disable")
      on Press: SetBit("ST_HMI_Var_HMI_bo_Disable")
      Appearance <- "ST_Main_Var_g_i16_Disable_Status"
   Button "OBJECT_108" at 873,370 size 177x68; TextOff '手动 / EXIT / 手動 / 수동'
      on Release: ResetBit("ST_HMI_Var_HMI_bo_Manual")
      on Press: SetBit("ST_HMI_Var_HMI_bo_Manual")
      Appearance <- "ST_Main_Var_g_i16_Manual_Status"
   Button "OBJECT_106" at 846,152 size 231x41; TextOff '手动 / EXIT / 手動 / 수동'; TextList "mode_enabled_4"
      ProcessValue <- "ST_Main_Var_g_i16_Mode_Enabled"
      Appearance <- "ST_Main_Var_g_i16_Mode_Enabled"
   Button "HmiScreenItemData_3" at 1119,386 size 159x47; TextOn '手动设置 / 手動設置 / 수동설정'; TextOff '动画 / 動画 / 애니메이션'
      on Release: ActivateScreen("动画", 0)
   Button "OBJECT_1" at 872,448 size 177x68; TextOff '回起点 EXIT 原点復帰 출발점으로 돌아가기'
      on Release: ResetBit("ST_HMI_Var_HMI_bo_Start_Position")
      on Press: SetBit("ST_HMI_Var_HMI_bo_Start_Position")
      Appearance <- "ST_Main_Var_g_i16_Mode_Enabled"
   Button "OBJECT_2" at 872,528 size 177x68; TextOff '启动 / EXIT / 起動 / 시작'
      on Release: ResetBit("ST_HMI_Var_HMI_bo_ZiDong_QiDong")
      on Press: SetBit("ST_HMI_Var_HMI_bo_ZiDong_QiDong")
      Appearance <- "ST_Main_Var_g_i16_Start_Position_Status"
   Button "OBJECT_3" at 40,536 size 177x68; TextOff 'SLM / EXIT'
      on Press: SetBit("ST_Main_Var_g_SLM_enable_status")
      Appearance <- "ST_Main_Var_g_SLM_enable_status"
   Button "OBJECT_4" at 40,616 size 177x68; TextOff '急停 / EXIT / 급정지'
      on Click: InvertBit("ST_Main_Var_g_bo_ZiDong_JiTing")
      Appearance <- "ST_Main_Var_g_bo_ZiDong_JiTing"
   TextField "Text Field_71" at 24,32 size 792x56; Text '手 动 控 制 / 手 動 制 御 / 수 동 제 어'
   TextField "Text Field_1" at 24,88 size 792x248; Text 'Text'
   Button "OBJECT_15" at 296,536 size 177x68; TextOff '电源通 / EXIT / 전원 on'
      Appearance <- "ST_Main_Var_g_bo_DI_1_D435_X122_2"
   Button "OBJECT_16" at 296,616 size 177x68; TextOff '电源断 / EXIT / 전원 off'
      on Release: ResetBit("ST_HMI_Var_HMI_bo_DianYuan_Duan")
      on Press: SetBit("ST_HMI_Var_HMI_bo_DianYuan_Duan")
   IOField "IO 域_20" at 873,219 size 176x41; Authorization "User administration"; FormatPattern 9
      on Activate: function_f41c6f6c("变量_1")
      ProcessValue <- "ST_Main_Var_g_i16_Manual_Status"
   Button "OBJECT_5" at 40,104 size 120x80; TextOff '出车 / EXIT / 出機 / 외진'
      on Release: ResetBit("ST_HMI_Var_HMI_bo_ChuChe")
      on Press: SetBit("ST_HMI_Var_HMI_bo_ChuChe")
      Appearance <- "ST_HMI_Var_HMI_bo_ChuChe"
   Button "OBJECT_7" at 200,104 size 120x80; TextOff '送条 / EXIT / 篠送り出し / 시누공급'
      on Release: InvertBit("ST_HMI_Var_HMI_bo_SongTiao")
      Appearance <- "ST_HMI_Var_HMI_bo_SongTiao"
   Button "OBJECT_9" at 360,104 size 120x80; TextOff '退绕 EXIT パッキン グオフ 언와인딩'
      on Release: ResetBit("ST_HMI_Var_HMI_bo_TuiRao")
      on Press: SetBit("ST_HMI_Var_HMI_bo_TuiRao")
      Appearance <- "ST_HMI_Var_HMI_bo_TuiRao"
   Button "OBJECT_12" at 520,104 size 120x80; TextOff '成形弓降 EXIT ワインデ ィング フォ ーラー下降 성형호랑 하강'
      on Release: ResetBit("ST_HMI_Var_HMI_bo_ChengXing_Down")
      on Press: SetBit("ST_HMI_Var_HMI_bo_ChengXing_Down")
      Appearance <- "ST_HMI_Var_HMI_bo_ChengXing_Down"
   Button "OBJECT_13" at 680,104 size 120x80; TextOff '张力弓升 EXIT カウンタ ーフォー ラー上昇 장력호랑 상승'
      on Release: ResetBit("ST_HMI_Var_HMI_bo_ZhangLi_Up")
      on Press: SetBit("ST_HMI_Var_HMI_bo_ZhangLi_Up")
      Appearance <- "ST_HMI_Var_HMI_bo_ZhangLi_Up"
   Button "OBJECT_6" at 40,232 size 120x80; TextOff '进车 / EXIT / 入機 / 내진'
      on Release: ResetBit("ST_HMI_Var_HMI_bo_JinChe")
      on Press: SetBit("ST_HMI_Var_HMI_bo_JinChe")
      Appearance <- "ST_HMI_Var_HMI_bo_JinChe"
   Button "OBJECT_8" at 200,232 size 120x80; TextOff '加捻 / EXIT / 撚掛 / 연사'
      on Release: ResetBit("ST_HMI_Var_HMI_bo_JiaNian")
      on Press: SetBit("ST_HMI_Var_HMI_bo_JiaNian")
      Appearance <- "ST_Main_Var_g_bo_JianNian_Jog_Status"
   Button "OBJECT_10" at 360,232 size 120x80; TextOff '卷绕 / EXIT / 巻取 / 와인딩'
      on Release: ResetBit("ST_HMI_Var_HMI_bo_JuanRao")
      on Press: SetBit("ST_HMI_Var_HMI_bo_JuanRao")
      Appearance <- "ST_HMI_Var_HMI_bo_JuanRao"
   Button "OBJECT_11" at 520,232 size 120x80; TextOff '成形弓升 EXIT ワインデ ィング フォ ーラー上昇 성형호랑 상승'
      on Release: ResetBit("ST_HMI_Var_HMI_bo_ChengXing_Up")
      on Press: SetBit("ST_HMI_Var_HMI_bo_ChengXing_Up")
      Appearance <- "ST_HMI_Var_HMI_bo_ChengXing_Up"
   Button "OBJECT_14" at 680,232 size 120x80; TextOff '张力弓降 EXIT カウンタ ーフォー ラー下降 장력호랑 하강'
      on Release: ResetBit("ST_HMI_Var_HMI_bo_ZhangLi_Down")
      on Press: SetBit("ST_HMI_Var_HMI_bo_ZhangLi_Down")
      Appearance <- "ST_HMI_Var_HMI_bo_ZhangLi_Down"